 2023 '~Spare WB2[63].7'; 2024 '~Spare WB2[63].8'; 2025 '~Spare WB2[63].9'; 2026 '~Spare WB2[63].10'; 2027 '~Spare WB2[63].11'; 2028 '~Spare WB2[63].12'; 2029 '~Spare WB2[63].13'; 2030 '~Spare WB2[63].14'; 2031 '~Spare WB2[63].15'; 2032 '~Spare WB2[63].16'; 2033 '~Spare WB2[63].17'; 2034 '~Spare WB2[63].18'; 2035 '~Spare WB2[63].19'; 2036 '~Spare WB2[63].20'; 2037 '~Spare WB2[63].21'; 2038 '~Spare WB2[63].22'; 2039 '~Spare WB2[63].23'; 2040 '~Spare WB2[63].24'; 2041 '~Spare WB2[63].25'; 2042 '~Spare WB2[63].26'; 2043 '~Spare WB2[63].27'; 2044 '~Spare WB2[63].28'; 2045 '~Spare WB2[63].29'; 2046 '~Spare WB2[63].30'; 2047 '~Spare WB2[63].31'; 2048 '~Spare WB2[64].0'; 2049 '~Spare WB2[64].1'; 2050 '~Spare WB2[64].2'; 2051 '~Spare WB2[64].3'; 2052 '~Spare WB2[64].4'; 2053 '~Spare WB2[64].5'; 2054 '~Spare WB2[64].6'; 2055 '~Spare WB2[64].7'; 2056 '~Spare WB2[64].8'; 2057 '~Spare WB2[64].9'; 2058 '~Spare WB2[64].10'; 2059 '~Spare WB2[64].11'; 2060 '~Spare WB2[64].12'; 2061 '~Spare WB2[64].13'; 2062 '~Spare WB2[64].14'; 2063 '~Spare WB2[64].15'; 2064 '~Spare WB2[64].16'; 2065 '~Spare WB2[64].17'; 2066 '~Spare WB2[64].18'; 2067 '~Spare WB2[64].19'; 2068 '~Spare WB2[64].20'; 2069 '~Spare WB2[64].21'; 2070 '~Spare WB2[64].22'; 2071 '~Spare WB2[64].23'; 2072 '~Spare WB2[64].24'; 2073 '~Spare WB2[64].25'; 2074 '~Spare WB2[64].26'; 2075 '~Spare WB2[64].27'; 2076 '~Spare WB2[64].28'; 2077 '~Spare WB2[64].29'; 2078 '~Spare WB2[64].30'; 2079 '~Spare WB2[64].31'; 2080 '~Spare WB2[65].0'; 2081 '~Spare WB2[65].1'; 2082 '~Spare WB2[65].2'; 2083 '~Spare WB2[65].3'; 2084 '~Spare WB2[65].4'; 2085 '~Spare WB2[65].5'; 2086 '~Spare WB2[65].6'; 2087 '~Spare WB2[65].7'; 2088 '~Spare WB2[65].8'; 2089 '~Spare WB2[65].9'; 2090 '~Spare WB2[65].10'; 2091 '~Spare WB2[65].11'; 2092 '~Spare WB2[65].12'; 2093 '~Spare WB2[65].13'; 2094 '~Spare WB2[65].14'; 2095 '~Spare WB2[65].15'; 2096 '~Spare WB2[65].16'; 2097 '~Spare WB2[65].17'; 2098 '~Spare WB2[65].18'; 2099 '~Spare WB2[65].19'; 2100 '~Spare WB2[65].20'; 2101 '~Spare WB2[65].21'; 2102 '~Spare WB2[65].22'; 2103 '~Spare WB2[65].23'; 2104 '~Spare WB2[65].24'; 2105 '~Spare WB2[65].25'; 2106 '~Spare WB2[65].26'; 2107 '~Spare WB2[65].27'; 2108 '~Spare WB2[65].28'; 2109 '~Spare WB2[65].29'; 2110 '~Spare WB2[65].30'; 2111 '~Spare WB2[65].31'; 2112 '~S001R16 Waiting Zone #1 Not Clear WB2[66].0'; 2113 '~S001R16 Waiting Zone #2 Not Clear WB2[66].1'; 2114 '~S001R16 Waiting Zone #3 Not Clear WB2[66].2'; 2115 '~S001R16 Waiting Zone #4 Not Clear WB2[66].3'; 2116 '~S001R16 Waiting Zone #5 Not Clear WB2[66].4'; 2117 '~S001R16 Waiting Zone #6 Not Clear WB2[66].5'; 2118 '~S001R16 Waiting Zone #7 Not Clear WB2[66].6'; 2119 '~S001R16 Waiting Zone #8 Not Clear WB2[66].7'; 2120 '~S001R16 Waiting Zone #9 Not Clear WB2[66].8'; 2121 '~S001R16 Waiting Zone #10 Not Clear WB2[66].9'; 2122 '~S001R16 Waiting Zone #11 Not Clear WB2[66].10'; 2123 '~S001R16 Waiting Zone #12 Not Clear WB2[66].11'; 2124 '~S001R16 Waiting Zone #13 Not Clear WB2[66].12'; 2125 '~S001R16 Waiting Zone #14 Not Clear WB2[66].13'; 2126 '~S001R16 Waiting Tip Dress Zone #1 Not Clear WB2[66].14'; 2127 '~S001R16 Waiting Tip Dress Zone #2 Not Clear WB2[66].15'; 2128 '~S001R16 Adjacent Robot xx-xx In Teach WB2[66].16'; 2129 '~S001R16 Adjacent Robot xx-xx In Teach WB2[66].17'; 2130 '~S001R16 Adjacent Robot xx-xx In Teach WB2[66].18'; 2131 '~S001R16 Adjacent Robot xx-xx In Teach WB2[66].19'; 2132 '~S001R16 Adjacent Robot xx-xx In Teach WB2[66].20'; 2133 '~S001R16 Adjacent Robot xx-xx In Teach WB2[66].21'; 2134 '~S001R16 Adjacent Robot xx-xx In Teach WB2[66].22'; 2135 '~S001R16 Adjacent Robot xx-xx In Teach WB2[66].23'; 2136 '~S001R16 Adjacent Robot xx-xx In Teach WB2[66].24'; 2137 '~S001R16 Adjacent Robot xx-xx In Teach WB2[66].25'; 2138 '~Spare WB2[66].26'; 2139 '~Spare WB2[66].27'; 2140 '~Spare WB2[66].28'; 2141 '~S001R16 Robot Not Clear Of Fixture WB2[66].29'; 2142 '~Spare WB2[66].30'; 2143 '~Spare WB2[66].31'; 2144 '~Spare WB2[67].0'; 2145 '~Spare WB2[67].1'; 2146 '~Spare WB2[67].2'; 2147 '~Spare WB2[67].3'; 2148 '~Spare WB2[67].4'; 2149 '~Spare WB2[67].5'; 2150 '~Spare WB2[67].6'; 2151 '~Spare WB2[67].7'; 2152 '~Spare WB2[67].8'; 2153 '~Spare WB2[67].9'; 2154 '~Spare WB2[67].10'; 2155 '~Spare WB2[67].11'; 2156 '~Spare WB2[67].12'; 2157 '~Spare WB2[67].13'; 2158 '~Spare WB2[67].14'; 2159 '~Spare WB2[67].15'; 2160 '~Spare WB2[67].16'; 2161 '~Spare WB2[67].17'; 2162 '~Spare WB2[67].18'; 2163 '~Spare WB2[67].19'; 2164 '~Spare WB2[67].20'; 2165 '~Spare WB2[67].21'; 2166 '~Spare WB2[67].22'; 2167 '~Spare WB2[67].23'; 2168 '~Spare WB2[67].24'; 2169 '~Spare WB2[67].25'; 2170 '~Spare WB2[67].26'; 2171 '~Spare WB2[67].27'; 2172 '~Spare WB2[67].28'; 2173 '~Spare WB2[67].29'; 2174 '~Spare WB2[67].30'; 2175 '~Spare WB2[67].31'; 2176 '~S001R16 Cycle Overtime WB2[68].0'; 2177 '~S001R16 In Bypass WB2[68].1'; 2178 '~S001R16 Battery Low WB2[68].2'; 2179 '~S001R16 Servo Over Torque WB2[68].3'; 2180 '~S001R16 Process Retry In Progress WB2[68].4'; 2181 '~Spare WB2[68].5'; 2182 '~S001R16 Robot Edit Occurred Ext App WB2[68].6'; 2183 '~S001R16 Robot Input Simmed WB2[68].7'; 2184 '~S001R16 Robot Output Simmed WB2[68].8'; 2185 '~Spare WB2[68].9'; 2186 '~Spare WB2[68].10'; 2187 '~Spare WB2[68].11'; 2188 '~Spare WB2[68].12'; 2189 '~Spare WB2[68].13'; 2190 '~Spare WB2[68].14'; 2191 '~Spare WB2[68].15'; 2192 '~S001R16F1B1.M.ModuleFlt - Externa App 1 I/O Module Warning WB2[68].16'; 2193 '~S001R16F2B1.M.ModuleFlt - Externa App 2 I/O Module Warning WB2[68].17'; 2194 '~S001R16F3B1.M.ModuleFlt - Externa App 3 I/O Module Warning WB2[68].18'; 2195 '~Spare WB2[68].19'; 2196 '~Spare WB2[68].20'; 2197 '~Spare WB2[68].21'; 2198 '~Spare WB2[68].22'; 2199 '~Spare WB2[68].23'; 2200 '~S001R16ES1 - S001R16 EtherNet Switch Port At Half Duplex WB2[68].24'; 2201 '~S001R16ES1 - S001R16 EtherNet Switch Config Changes Not Saved WB2[68].25'; 2202 '~S001R16ES1 - S001R16 EtherNet Switch Configuration Changed WB2[68].26'; 2203 '~S001R16ES1 - S001R16 EtherNet Switch Port With Excessive Errors WB2[68].27'; 2204 '~S001R16ES1 - S001R16 EtherNet Switch Port With Utilization Warning WB2[68].28'; 2205 '~S001R16ES1 - S001R16 EtherNet Switch Changes Require Reboot WB2[68].29'; 2206 '~Spare WB2[68].30'; 2207 '~Spare WB2[68].31'; 2208 '~Spare WB2[69].0'; 2209 '~Spare WB2[69].1'; 2210 '~S001R16 Servo Gun Tip Calib Request 1 WB2[69].2'; 2211 '~S001R16 I-Available Warning 1 WB2[69].3'; 2212 '~S001R16 Tip Dress Motor 1 Fault Bypassed WB2[69].4'; 2213 '~S001R16 Tip Change Notice 1 WB2[69].5'; 2214 '~S001R16 Bypass Tip Dresser 1 Selected WB2[69].6'; 2215 '~S001R16 Auto Tip Changer Low 1 WB2[69].7'; 2216 '~S001R16 Auto Tip Changer Empty 1 WB2[69].8'; 2217 '~S001R16 Tip Wear Ratio Warning 1 - Touch Up Tip Dress Program WB2[69].9'; 2218 '~S001R16 Stud Weld 1 Maintenance Reqd WB2[69].10'; 2219 '~S001R16 Stud Weld 1 Low Stud Warning WB2[69].11'; 2220 '~Spare WB2[69].12'; 2221 '~S001R16 Rivet 1 Low Rivet Warning WB2[69].13'; 2222 '~S001R16 Rivet 1 - Skip Once Initiated from Robot TP WB2[69].14'; 2223 '~S001R16 Rivet 1 - Skip Remaining Initiated from Robot TP WB2[69].15'; 2224 '~S001R16 Rivet 1 Preventive Maintenace Required WB2[69].16'; 2225 '~S001R16 Rivet 1 Magazine Low WB2[69].17'; 2226 '~S001R16 Tip Change 1 Bypassed WB2[69].18'; 2227 '~S001R16 Mig Weld Fluid Level Low WB2[69].19'; 2228 '~S001R16 Weld Ctrlr 1 Adaptive Mode Is Disabled WB2[69].20'; 2229 '~S001R16 Tip Cutter 1 Warning WB2[69].21'; 2230 '~S001R16 Rivet 1 Tape-Cut Required WB2[69].22'; 2231 '~S001R16 Wire Feeder Motor Over Current WB2[69].23'; 2232 '~Spare WB2[69].24'; 2233 '~S001R16 Sealer Ctrlr 1 Minor Fault WB2[69].25'; 2234 '~S001R16 Sealer Ctrlr 1 Required Rezeroing WB2[69].26'; 2235 '~S001R16 Loaded To Average WB2[69].27'; 2236 '~S001R16 Vision Process Aborted WB2[69].28'; 2237 '~S001R16 Vision System Trending WB2[69].29'; 2238 '~S001R16 Vision Out Of Tolerance WB2[69].30'; 2239 '~Spare WB2[69].31'; 2240 '~Spare WB2[70].0'; 2241 '~Spare WB2[70].1'; 2242 '~S001R16 Servo Gun Tip Calib Request 2 WB2[70].2'; 2243 '~S001R16 I-Available Warning 2 WB2[70].3'; 2244 '~S001R16 Tip Dress Motor 2 Fault Bypassed WB2[70].4'; 2245 '~S001R16 Tip Change Notice 2 WB2[70].5'; 2246 '~S001R16 Bypass Tip Dresser 2 Selected WB2[70].6'; 2247 '~S001R16 Auto Tip Changer Low 2 WB2[70].7'; 2248 '~S001R16 Auto Tip Changer Empty 2 WB2[70].8'; 2249 '~S001R16 Tip Wear Ratio Warning 2 - Touch Up Tip Dress Program WB2[70].9'; 2250 '~S001R16 Stud Weld 2 Maintenance Reqd WB2[70].10'; 2251 '~S001R16 Stud Weld 2 Low Stud Warning WB2[70].11'; 2252 '~Spare WB2[70].12'; 2253 '~S001R16 Rivet 2 Low Rivet Warning WB2[70].13'; 2254 '~S001R16 Rivet 2 - Skip Once Initiated from Robot TP WB2[70].14'; 2255 '~S001R16 Rivet 2 - Skip Remaining Initiated from Robot TP WB2[70].15'; 2256 '~S001R16 Rivet 2 Preventive Maintenace Required WB2[70].16'; 2257 '~S001R16 Rivet 2 Magazine Low WB2[70].17'; 2258 '~S001R16 Tip Change 2 Bypassed WB2[70].18'; 2259 '~S001R16 Laser Dirty Glass Warning WB2[70].19'; 2260 '~S001R16 Weld Ctrlr 2 Adaptive Mode Is Disabled WB2[70].20'; 2261 '~S001R16 Tip Cutter 2 Warning WB2[70].21'; 2262 '~S001R16 Rivet 2 Tape-Cut Required WB2[70].22'; 2263 '~S001R16 Mig Tip Nozzel Replacement Warning WB2[70].23'; 2264 '~S001R16 Mig Tip Nozzel Replacement Required WB2[70].24'; 2265 '~S001R16 Sealer Ctrlr 2 Minor Fault WB2[70].25'; 2266 '~S001R16 Sealer Ctrlr 2 Required Rezeroing WB2[70].26'; 2267 '~S001R16 Mig Barrel Replacement Warning WB2[70].27'; 2268 '~S001R16 Mig Barrel Replacement Required WB2[70].28'; 2269 '~S001R16 In Touch Up Mode WB2[70].29'; 2270 '~S001R16 Touch Up Mode Not Enabled WB2[70].30'; 2271 '~Spare WB2[70].31'; 2272 '~S001R16 Laser Controller Fault WB2[71].0'; 2273 '~S001R16 Laser Dirty Glass Warning WB2[71].1'; 2274 '~S001R16 Laser Warning WB2[71].2'; 2275 '~Spare WB2[71].3'; 2276 '~Spare WB2[71].4'; 2277 '~Spare WB2[71].5'; 2278 '~Spare WB2[71].6'; 2279 '~Spare WB2[71].7'; 2280 '~Spare WB2[71].8'; 2281 '~Spare WB2[71].9'; 2282 '~Spare WB2[71].10'; 2283 '~Spare WB2[71].11'; 2284 '~Spare WB2[71].12'; 2285 '~Spare WB2[71].13'; 2286 '~Spare WB2[71].14'; 2287 '~Spare WB2[71].15'; 2288 '~Spare WB2[71].16'; 2289 '~Spare WB2[71].17'; 2290 '~Spare WB2[71].18'; 2291 '~Spare WB2[71].19'; 2292 '~Spare WB2[71].20'; 2293 '~Spare WB2[71].21'; 2294 '~Spare WB2[71].22'; 2295 '~Spare WB2[71].23'; 2296 '~Spare WB2[71].24'; 2297 '~Spare WB2[71].25'; 2298 '~Spare WB2[71].26'; 2299 '~Spare WB2[71].27'; 2300 '~Spare WB2[71].28'; 2301 '~Spare WB2[71].29'; 2302 '~Spare WB2[71].30'; 2303 '~Spare WB2[71].31'; 2304 '~Spare WB2[72].0'; 2305 '~Spare WB2[72].1'; 2306 '~Spare WB2[72].2'; 2307 '~Spare WB2[72].3'; 2308 '~Spare WB2[72].4'; 2309 '~Spare WB2[72].5'; 2310 '~Spare WB2[72].6'; 2311 '~Spare WB2[72].7'; 2312 '~Spare WB2[72].8'; 2313 '~Spare WB2[72].9'; 2314 '~Spare WB2[72].10'; 2315 '~Spare WB2[72].11'; 2316 '~Spare WB2[72].12'; 2317 '~Spare WB2[72].13'; 2318 '~Spare WB2[72].14'; 2319 '~Spare WB2[72].15'; 2320 '~Spare WB2[72].16'; 2321 '~Spare WB2[72].17'; 2322 '~Spare WB2[72].18'; 2323 '~Spare WB2[72].19'; 2324 '~Spare WB2[72].20'; 2325 '~Spare WB2[72].21'; 2326 '~Spare WB2[72].22'; 2327 '~Spare WB2[72].23'; 2328 '~Spare WB2[72].24'; 2329 '~Spare WB2[72].25'; 2330 '~Spare WB2[72].26'; 2331 '~Spare WB2[72].27'; 2332 '~Spare WB2[72].28'; 2333 '~Spare WB2[72].29'; 2334 '~Spare WB2[72].30'; 2335 '~Spare WB2[72].31'; 2336 '~Spare WB2[73].0'; 2337 '~Spare WB2[73].1'; 2338 '~Spare WB2[73].2'; 2339 '~Spare WB2[73].3'; 2340 '~Spare WB2[73].4'; 2341 '~Spare WB2[73].5'; 2342 '~Spare WB2[73].6'; 2343 '~Spare WB2[73].7'; 2344 '~Spare WB2[73].8'; 2345 '~Spare WB2[73].9'; 2346 '~Spare WB2[73].10'; 2347 '~Spare WB2[73].11'; 2348 '~Spare WB2[73].12'; 2349 '~Spare WB2[73].13'; 2350 '~Spare WB2[73].14'; 2351 '~Spare WB2[73].15'; 2352 '~Spare WB2[73].16'; 2353 '~Spare WB2[73].17'; 2354 '~Spare WB2[73].18'; 2355 '~Spare WB2[73].19'; 2356 '~Spare WB2[73].20'; 2357 '~Spare WB2[73].21'; 2358 '~Spare WB2[73].22'; 2359 '~Spare WB2[73].23'; 2360 '~Spare WB2[73].24'; 2361 '~Spare WB2[73].25'; 2362 '~Spare WB2[73].26'; 2363 '~Spare WB2[73].27'; 2364 '~Spare WB2[73].28'; 2365 '~Spare WB2[73].29'; 2366 '~Spare WB2[73].30'; 2367 '~Spare WB2[73].31'; 2368 '~Spare WB2[74].0'; 2369 '~Spare WB2[74].1'; 2370 '~Spare WB2[74].2'; 2371 '~Spare WB2[74].3'; 2372 '~Spare WB2[74].4'; 2373 '~Spare WB2[74].5'; 2374 '~Spare WB2[74].6'; 2375 '~Spare WB2[74].7'; 2376 '~Spare WB2[74].8'; 2377 '~Spare WB2[74].9'; 2378 '~Spare WB2[74].10'; 2379 '~Spare WB2[74].11'; 2380 '~Spare WB2[74].12'; 2381 '~Spare WB2[74].13'; 2382 '~Spare WB2[74].14'; 2383 '~Spare WB2[74].15'; 2384 '~Spare WB2[74].16'; 2385 '~Spare WB2[74].17'; 2386 '~Spare WB2[74].18'; 2387 '~Spare WB2[74].19'; 2388 '~Spare WB2[74].20'; 2389 '~Spare WB2[74].21'; 2390 '~Spare WB2[74].22'; 2391 '~Spare WB2[74].23'; 2392 '~Spare WB2[74].24'; 2393 '~Spare WB2[74].25'; 2394 '~Spare WB2[74].26'; 2395 '~Spare WB2[74].27'; 2396 '~Spare WB2[74].28'; 2397 '~Spare WB2[74].29'; 2398 '~Spare WB2[74].30'; 2399 '~Spare WB2[74].31'; 2400 '~S002 Fixture Cycle Over Time WB2[75].0'; 2401 '~S002CV1 Conveyor Over Cycle Time WB2[75].1'; 2402 '~Spare WB2[75].2'; 2403 '~Spare WB2[75].3'; 2404 '~S002CV1 ~ Conveyor Drive Brake Still Released WB2[75].4'; 2405 '~Spare WB2[75].5'; 2406 '~Spare WB2[75].6'; 2407 '~Spare WB2[75].7'; 2408 '~Spare WB2[75].8'; 2409 '~Spare WB2[75].9'; 2410 '~S002CV1DES1 - S002CV1 EtherNet Switch Port At Half Duplex WB2[75].10'; 2411 '~S002CV1DES1 - S002CV1 EtherNet Switch Config Changes Not Saved WB2[75].11'; 2412 '~S002CV1DES1 - S002CV1 EtherNet Switch Configuration Changed WB2[75].12'; 2413 '~S002CV1DES1 - S002CV1 EtherNet Switch Port With Excessive Errors WB2[75].13'; 2414 '~S002CV1DES1 - S002CV1 EtherNet Switch Port With Utilization Warn WB2[75].14'; 2415 '~S002CV1DES1 - S002CV1 EtherNet Switch Changes Require Reboot WB2[75].15'; 2416 '~Spare WB2[75].16'; 2417 '~Spare WB2[75].17'; 2418 '~Spare WB2[75].18'; 2419 '~Spare WB2[75].19'; 2420 '~Spare WB2[75].20'; 2421 '~Spare WB2[75].21'; 2422 '~Spare WB2[75].22'; 2423 '~Spare WB2[75].23'; 2424 '~Spare WB2[75].24'; 2425 '~Spare WB2[75].25'; 2426 '~Spare WB2[75].26'; 2427 '~Spare WB2[75].27'; 2428 '~Spare WB2[75].28'; 2429 '~Spare WB2[75].29'; 2430 '~Spare WB2[75].30'; 2431 '~Spare WB2[75].31'; 2432 '~S002WC# Tip Change Required Warning WB2[76].0'; 2433 '~S002WC# Tip Change Required Warning WB2[76].1'; 2434 '~S002WC# Tip Change Required Warning WB2[76].2'; 2435 '~S002WC# Tip Change Required Warning WB2[76].3'; 2436 '~S002WC# Tip Change Required Warning WB2[76].4'; 2437 '~S002WC# Tip Change Required Warning WB2[76].5'; 2438 '~Spare WB2[76].6'; 2439 '~S003TL1DES1 - S003TL1 EtherNet Switch Port At Half Duplex WB2[76].7'; 2440 '~S003TL1DES1 - S003TL1 EtherNet Switch Config Changes Not Saved WB2[76].8'; 2441 '~S003TL1DES1 - S003TL1 EtherNet Switch Configuration Changed WB2[76].9'; 2442 '~S003TL1DES1 - S003TL1 EtherNet Switch Port With Excessive Errors WB2[76].10'; 2443 '~S003TL1DES1 - S003TL1 EtherNet Switch Port With Utilization Warn WB2[76].11'; 2444 '~S003TL1DES1 - S003TL1 EtherNet Switch Changes Require Reboot WB2[76].12'; 2445 '~Spare WB2[76].13'; 2446 '~Spare WB2[76].14'; 2447 '~Spare WB2[76].15'; 2448 '~S003TL1 Turn Table Index Over Cycle Time WB2[76].16'; 2449 '~S003TL1 Tool-Tray VFD Drive Temperature Warning WB2[76].17'; 2450 '~S003TL1 Fixture A Bypassed WB2[76].18'; 2451 '~S003TL1 Fixture B Bypassed WB2[76].19'; 2452 '~S003TL1 Fixture C Bypassed WB2[76].20'; 2453 '~Spare WB2[76].21'; 2454 '~S003TL1 Major Motion Not Enabled WB2[76].22'; 2455 '~S003TL1 All Robots Not Clear Of Turn Table WB2[76].23'; 2456 '~S003TL1 All Tooling Not Clear To Rotate WB2[76].24'; 2457 '~S003TL1 Light Screen Not Clear For Rotate WB2[76].25'; 2458 '~S003TL1 Tool Tray Brake Still Released WB2[76].26'; 2459 '~Spare WB2[76].27'; 2460 '~Spare WB2[76].28'; 2461 '~Spare WB2[76].29'; 2462 '~Spare WB2[76].30'; 2463 '~Spare WB2[76].31'; 2464 '~Spare WB2[77].0'; 2465 '~Spare WB2[77].1'; 2466 '~Spare WB2[77].2'; 2467 '~Spare WB2[77].3'; 2468 '~Spare WB2[77].4'; 2469 '~Spare WB2[77].5'; 2470 '~Spare WB2[77].6'; 2471 '~Spare WB2[77].7'; 2472 '~Spare WB2[77].8'; 2473 '~Spare WB2[77].9'; 2474 '~Spare WB2[77].10'; 2475 '~Spare WB2[77].11'; 2476 '~Spare WB2[77].12'; 2477 '~Spare WB2[77].13'; 2478 '~Spare WB2[77].14'; 2479 '~Spare WB2[77].15'; 2480 '~Spare WB2[77].16'; 2481 '~Spare WB2[77].17'; 2482 '~Spare WB2[77].18'; 2483 '~Spare WB2[77].19'; 2484 '~Spare WB2[77].20'; 2485 '~Spare WB2[77].21'; 2486 '~Spare WB2[77].22'; 2487 '~Spare WB2[77].23'; 2488 '~Spare WB2[77].24'; 2489 '~Spare WB2[77].25'; 2490 '~Spare WB2[77].26'; 2491 '~Spare WB2[77].27'; 2492 '~Spare WB2[77].28'; 2493 '~Spare WB2[77].29'; 2494 '~Spare WB2[77].30'; 2495 '~Spare WB2[77].31'; 2496 '~Spare WB2[78].0'; 2497 '~S001CV1 Conveyor Over Cycle Time WB2[78].1'; 2498 '~S001CV1 Conveyor Auto/Mastering SS in Mastering Position WB2[78].2'; 2499 '~S001CV1 Operator Over Cycle Time WB2[78].3'; 2500 '~S001CV1 Conveyor Part Low Level Warning WB2[78].4'; 2501 '~S001CV1 ~ Conveyor Drive Brake Still Released WB2[78].5'; 2502 '~Spare WB2[78].6'; 2503 '~Spare WB2[78].7'; 2504 '~Spare WB2[78].8'; 2505 '~Spare WB2[78].9'; 2506 '~S001CV1DES1 - S001CV1 EtherNet Switch Port At Half Duplex WB2[78].10'; 2507 '~S001CV1DES1 - S001CV1 EtherNet Switch Config Changes Not Saved WB2[78].11'; 2508 '~S001CV1DES1 - S001CV1 EtherNet Switch Configuration Changed WB2[78].12'; 2509 '~S001CV1DES1 - S001CV1 EtherNet Switch Port With Excessive Errors WB2[78].13'; 2510 '~S001CV1DES1 - S001CV1 EtherNet Switch Port With Utilization Warn WB2[78].14'; 2511 '~S001CV1DES1 - S001CV1 EtherNet Switch Changes Require Reboot WB2[78].15'; 2512 '~Spare WB2[78].16'; 2513 '~Spare WB2[78].17'; 2514 '~Spare WB2[78].18'; 2515 '~Spare WB2[78].19'; 2516 '~Spare WB2[78].20'; 2517 '~Spare WB2[78].21'; 2518 '~Spare WB2[78].22'; 2519 '~Spare WB2[78].23'; 2520 '~Spare WB2[78].24'; 2521 '~Spare WB2[78].25'; 2522 '~Spare WB2[78].26'; 2523 '~Spare WB2[78].27'; 2524 '~Spare WB2[78].28'; 2525 '~Spare WB2[78].29'; 2526 '~Spare WB2[78].30'; 2527 '~Spare WB2[78].31'; 2528 '~S001TT1 Operator Load Cycle Overtime WB2[79].0'; 2529 '~S001TT1 Index Cycle Overtime WB2[79].1'; 2530 '~Spare WB2[79].2'; 2531 '~Spare WB2[79].3'; 2532 '~S001TT1 VFD Temperature Warning WB2[79].4'; 2533 '~S001TT1 Turn Table Brake Still Released WB2[79].5'; 2534 '~Spare WB2[79].6'; 2535 '~Spare WB2[79].7'; 2536 '~S001TT1 Fixture A Bypass Selected WB2[79].8'; 2537 '~S001TT1 Fixture B Bypass Selected WB2[79].9'; 2538 '~S001TT1 Fixture C Bypass Selected WB2[79].10'; 2539 '~S001TT1 Fixture D Bypass Selected WB2[79].11'; 2540 '~Spare WB2[79].12'; 2541 '~S001TT1 Manual Mode Motion Not Enabled WB2[79].13'; 2542 '~S001TT1 Lt Screen Not Clear Or Active WB2[79].14'; 2543 '~S001TT1 Robots Not Clear Of Turntable Index WB2[79].15'; 2544 '~S001TT1 All Tooling Not Clear To Rotate WB2[79].16'; 2545 '~Spare WB2[79].17'; 2546 '~S001TT1DES1 - S001TT1 EtherNet Switch Port At Half Duplex WB2[79].18'; 2547 '~S001TT1DES1 - S001TT1 EtherNet Switch Config Changes Not Saved WB2[79].19'; 2548 '~S001TT1DES1 - S001TT1 EtherNet Switch Configuration Changed WB2[79].20'; 2549 '~S001TT1DES1 - S001TT1 EtherNet Switch Port With Excessive Errors WB2[79].21'; 2550 '~S001TT1DES1 - S001TT1 EtherNet Switch Port With Utilization Warn WB2[79].22'; 2551 '~S001TT1DES1 - S001TT1 EtherNet Switch Changes Require Reboot WB2[79].23'; 2552 '~Spare WB2[79].24'; 2553 '~S001TT1DES2 - S001TT1 EtherNet Switch Port At Half Duplex WB2[79].25'; 2554 '~S001TT1DES2 - S001TT1 EtherNet Switch Config Changes Not Saved WB2[79].26'; 2555 '~S001TT1DES2 - S001TT1 EtherNet Switch Configuration Changed WB2[79].27'; 2556 '~S001TT1DES2 - S001TT1 EtherNet Switch Port With Excessive Errors WB2[79].28'; 2557 '~S001TT1DES2 - S001TT1 EtherNet Switch Port With Utilization Warn WB2[79].29'; 2558 '~S001TT1DES2 - S001TT1 EtherNet Switch Changes Require Reboot WB2[79].30'; 2559 '~Spare WB2[79].31'; 2560 '~S002TT1 Operator Load Cycle Overtime WB2[80].0'; 2561 '~S002TT1 Index Cycle Overtime WB2[80].1'; 2562 '~Spare 